(* Logix 5000 project; controller FV vendor 1 type 14 code 217 rev 31.11; software revision 31.00; part 60 of 63 *)
(* tags used below, declared in another part *)
   YP_B103 : INT[15];   // Original N File From SLC, No Description Available
   YP_B103_1_1_Storagebit : BOOL;
   YP_B30 : INT[37];   // Original N File From SLC, No Description Available
   YP_B31 : INT[37];   // Original N File From SLC, No Description Available
   YP_B92 : INT[105];   // Original N File From SLC, No Description Available
   YP_N32 : INT[257];
   YP_N55 : INT[244];   // Original N File From SLC, No Description Available
   YP_N7 : INT[56];   // INTEGER
   YP_SYSTEM_4_BIT6_TIMEBASE : ALIAS FOR One_Second_1_scan;
(* YP_Common, continued *)

   47: [AND(YP_B92[4],YP_B92[44],YP_B92[44]) ,OR(YP_B92[4],YP_B92[24],YP_B92[64]) ,XOR(YP_B92[44],YP_B92[64],YP_B92[24]) ];
   48: [AND(YP_B92[5],YP_B92[45],YP_B92[45]) ,OR(YP_B92[5],YP_B92[25],YP_B92[65]) ,XOR(YP_B92[45],YP_B92[65],YP_B92[25]) ];
   49: [AND(YP_B92[6],YP_B92[46],YP_B92[46]) ,OR(YP_B92[6],YP_B92[26],YP_B92[66]) ,XOR(YP_B92[46],YP_B92[66],YP_B92[26]) ];
   50: [AND(YP_B92[7],YP_B92[47],YP_B92[47]) ,OR(YP_B92[7],YP_B92[27],YP_B92[67]) ,XOR(YP_B92[47],YP_B92[67],YP_B92[27]) ];
   51: [AND(YP_B92[8],YP_B92[48],YP_B92[48]) ,OR(YP_B92[8],YP_B92[28],YP_B92[68]) ,XOR(YP_B92[48],YP_B92[68],YP_B92[28]) ];
   52: [AND(YP_B92[9],YP_B92[49],YP_B92[49]) ,OR(YP_B92[9],YP_B92[29],YP_B92[69]) ,XOR(YP_B92[49],YP_B92[69],YP_B92[29]) ];
   53: [AND(YP_B92[10],YP_B92[50],YP_B92[50]) ,OR(YP_B92[10],YP_B92[30],YP_B92[70]) ,XOR(YP_B92[50],YP_B92[70],YP_B92[30]) ];
   54: [AND(YP_B92[11],YP_B92[51],YP_B92[51]) ,OR(YP_B92[11],YP_B92[31],YP_B92[71]) ,XOR(YP_B92[51],YP_B92[71],YP_B92[31]) ];
   55: [AND(YP_B92[12],YP_B92[52],YP_B92[52]) ,OR(YP_B92[12],YP_B92[32],YP_B92[72]) ,XOR(YP_B92[52],YP_B92[72],YP_B92[32]) ];
   56: [AND(YP_B92[13],YP_B92[53],YP_B92[53]) ,OR(YP_B92[13],YP_B92[33],YP_B92[73]) ,XOR(YP_B92[53],YP_B92[73],YP_B92[33]) ];
   57: [AND(YP_B92[14],YP_B92[54],YP_B92[54]) ,OR(YP_B92[14],YP_B92[34],YP_B92[74]) ,XOR(YP_B92[54],YP_B92[74],YP_B92[34]) ];
   58: [AND(YP_B92[15],YP_B92[55],YP_B92[55]) ,OR(YP_B92[15],YP_B92[35],YP_B92[75]) ,XOR(YP_B92[55],YP_B92[75],YP_B92[35]) ];
   59: [AND(YP_B92[16],YP_B92[56],YP_B92[56]) ,OR(YP_B92[16],YP_B92[36],YP_B92[76]) ,XOR(YP_B92[56],YP_B92[76],YP_B92[36]) ];
   60: [AND(YP_B92[17],YP_B92[57],YP_B92[57]) ,OR(YP_B92[17],YP_B92[37],YP_B92[77]) ,XOR(YP_B92[57],YP_B92[77],YP_B92[37]) ];
   61: [AND(YP_B92[18],YP_B92[58],YP_B92[58]) ,OR(YP_B92[18],YP_B92[38],YP_B92[78]) ,XOR(YP_B92[58],YP_B92[78],YP_B92[38]) ];
   62: [AND(YP_B92[19],YP_B92[59],YP_B92[59]) ,OR(YP_B92[19],YP_B92[39],YP_B92[79]) ,XOR(YP_B92[59],YP_B92[79],YP_B92[39]) ];
   63: [XIC(YP_B30[31].4) ,XIC(YP_B103[1].2) ]OSR(YP_B103[1].1,YP_B103_1_1_Storagebit)XIC(YP_B103_1_1_Storagebit)OTE(YP_B103[1].0);
   64: XIC(YP_B103[1].2)OTU(YP_B103[1].2);
   65: XIC(YP_B103[1].0)[OR(YP_B92[20],YP_B92[40],YP_B92[40]) ,AND(YP_B92[0],YP_B92[20],YP_B92[20]) ];
   66: XIC(YP_B103[1].0)[OR(YP_B92[21],YP_B92[41],YP_B92[41]) ,AND(YP_B92[1],YP_B92[21],YP_B92[21]) ];
   67: XIC(YP_B103[1].0)[OR(YP_B92[22],YP_B92[42],YP_B92[42]) ,AND(YP_B92[2],YP_B92[22],YP_B92[22]) ];
   68: XIC(YP_B103[1].0)[OR(YP_B92[23],YP_B92[43],YP_B92[43]) ,AND(YP_B92[3],YP_B92[23],YP_B92[23]) ];
   69: XIC(YP_B103[1].0)[OR(YP_B92[24],YP_B92[44],YP_B92[44]) ,AND(YP_B92[4],YP_B92[24],YP_B92[24]) ];
   70: XIC(YP_B103[1].0)[OR(YP_B92[25],YP_B92[45],YP_B92[45]) ,AND(YP_B92[5],YP_B92[25],YP_B92[25]) ];
   71: XIC(YP_B103[1].0)[OR(YP_B92[26],YP_B92[46],YP_B92[46]) ,AND(YP_B92[6],YP_B92[26],YP_B92[26]) ];
   72: XIC(YP_B103[1].0)[OR(YP_B92[27],YP_B92[47],YP_B92[47]) ,AND(YP_B92[7],YP_B92[27],YP_B92[27]) ];
   73: XIC(YP_B103[1].0)[OR(YP_B92[28],YP_B92[48],YP_B92[48]) ,AND(YP_B92[8],YP_B92[28],YP_B92[28]) ];
   74: XIC(YP_B103[1].0)[OR(YP_B92[29],YP_B92[49],YP_B92[49]) ,AND(YP_B92[9],YP_B92[29],YP_B92[29]) ];
   75: XIC(YP_B103[1].0)[OR(YP_B92[30],YP_B92[50],YP_B92[50]) ,AND(YP_B92[10],YP_B92[30],YP_B92[30]) ];
   76: XIC(YP_B103[1].0)[OR(YP_B92[31],YP_B92[51],YP_B92[51]) ,AND(YP_B92[11],YP_B92[31],YP_B92[31]) ];
   77: XIC(YP_B103[1].0)[OR(YP_B92[32],YP_B92[52],YP_B92[52]) ,AND(YP_B92[12],YP_B92[32],YP_B92[32]) ];
   78: XIC(YP_B103[1].0)[OR(YP_B92[33],YP_B92[53],YP_B92[53]) ,AND(YP_B92[13],YP_B92[33],YP_B92[33]) ];
   79: XIC(YP_B103[1].0)[OR(YP_B92[34],YP_B92[54],YP_B92[54]) ,AND(YP_B92[14],YP_B92[34],YP_B92[34]) ];
   80: XIC(YP_B103[1].0)[OR(YP_B92[35],YP_B92[55],YP_B92[55]) ,AND(YP_B92[15],YP_B92[35],YP_B92[35]) ];
   81: XIC(YP_B103[1].0)[OR(YP_B92[36],YP_B92[56],YP_B92[56]) ,AND(YP_B92[16],YP_B92[36],YP_B92[36]) ];
   82: XIC(YP_B103[1].0)[OR(YP_B92[37],YP_B92[57],YP_B92[57]) ,AND(YP_B92[17],YP_B92[37],YP_B92[37]) ];
   83: XIC(YP_B103[1].0)[OR(YP_B92[38],YP_B92[58],YP_B92[58]) ,AND(YP_B92[18],YP_B92[38],YP_B92[38]) ];
   84: XIC(YP_B103[1].0)[OR(YP_B92[39],YP_B92[59],YP_B92[59]) ,AND(YP_B92[19],YP_B92[39],YP_B92[39]) ];
   85: XIC(YP_B103[1].0)MOV(0,YP_N7[38]);
   86: XIC(YP_SYSTEM_4_BIT6_TIMEBASE)MOV(YP_B92[60],YP_B92[80]);
   87: XIO(YP_SYSTEM_4_BIT6_TIMEBASE)MOV(YP_B92[40],YP_B92[80]);
   88: XIC(YP_SYSTEM_4_BIT6_TIMEBASE)MOV(YP_B92[61],YP_B92[81]);
   89: XIO(YP_SYSTEM_4_BIT6_TIMEBASE)MOV(YP_B92[41],YP_B92[81]);
   90: XIC(YP_SYSTEM_4_BIT6_TIMEBASE)MOV(YP_B92[62],YP_B92[82]);
   91: XIO(YP_SYSTEM_4_BIT6_TIMEBASE)MOV(YP_B92[42],YP_B92[82]);
   92: XIC(YP_SYSTEM_4_BIT6_TIMEBASE)MOV(YP_B92[63],YP_B92[83]);
   93: XIO(YP_SYSTEM_4_BIT6_TIMEBASE)MOV(YP_B92[43],YP_B92[83]);
   94: XIC(YP_SYSTEM_4_BIT6_TIMEBASE)MOV(YP_B92[64],YP_B92[84]);
   95: XIO(YP_SYSTEM_4_BIT6_TIMEBASE)MOV(YP_B92[44],YP_B92[84]);
   96: XIC(YP_SYSTEM_4_BIT6_TIMEBASE)MOV(YP_B92[65],YP_B92[85]);
   97: XIO(YP_SYSTEM_4_BIT6_TIMEBASE)MOV(YP_B92[45],YP_B92[85]);
   98: XIC(YP_SYSTEM_4_BIT6_TIMEBASE)MOV(YP_B92[66],YP_B92[86]);
   99: XIO(YP_SYSTEM_4_BIT6_TIMEBASE)MOV(YP_B92[46],YP_B92[86]);
   100: XIC(YP_SYSTEM_4_BIT6_TIMEBASE)MOV(YP_B92[67],YP_B92[87]);
   101: XIO(YP_SYSTEM_4_BIT6_TIMEBASE)MOV(YP_B92[47],YP_B92[87]);
   102: XIC(YP_SYSTEM_4_BIT6_TIMEBASE)MOV(YP_B92[68],YP_B92[88]);
   103: XIO(YP_SYSTEM_4_BIT6_TIMEBASE)MOV(YP_B92[48],YP_B92[88]);
   104: XIC(YP_SYSTEM_4_BIT6_TIMEBASE)MOV(YP_B92[69],YP_B92[89]);
   105: XIO(YP_SYSTEM_4_BIT6_TIMEBASE)MOV(YP_B92[49],YP_B92[89]);
   106: XIC(YP_SYSTEM_4_BIT6_TIMEBASE)MOV(YP_B92[70],YP_B92[90]);
   107: XIO(YP_SYSTEM_4_BIT6_TIMEBASE)MOV(YP_B92[50],YP_B92[90]);
   108: XIC(YP_SYSTEM_4_BIT6_TIMEBASE)MOV(YP_B92[71],YP_B92[91]);
   109: XIO(YP_SYSTEM_4_BIT6_TIMEBASE)MOV(YP_B92[51],YP_B92[91]);
   110: XIC(YP_SYSTEM_4_BIT6_TIMEBASE)MOV(YP_B92[72],YP_B92[92]);
   111: XIO(YP_SYSTEM_4_BIT6_TIMEBASE)MOV(YP_B92[52],YP_B92[92]);
   112: XIC(YP_SYSTEM_4_BIT6_TIMEBASE)MOV(YP_B92[73],YP_B92[93]);
   113: XIO(YP_SYSTEM_4_BIT6_TIMEBASE)MOV(YP_B92[53],YP_B92[93]);
   114: XIC(YP_SYSTEM_4_BIT6_TIMEBASE)MOV(YP_B92[74],YP_B92[94]);
   115: XIO(YP_SYSTEM_4_BIT6_TIMEBASE)MOV(YP_B92[54],YP_B92[94]);
   116: XIC(YP_SYSTEM_4_BIT6_TIMEBASE)MOV(YP_B92[75],YP_B92[95]);
   117: XIO(YP_SYSTEM_4_BIT6_TIMEBASE)MOV(YP_B92[55],YP_B92[95]);
   118: XIC(YP_SYSTEM_4_BIT6_TIMEBASE)MOV(YP_B92[76],YP_B92[96]);
   119: XIO(YP_SYSTEM_4_BIT6_TIMEBASE)MOV(YP_B92[56],YP_B92[96]);
   120: XIC(YP_SYSTEM_4_BIT6_TIMEBASE)MOV(YP_B92[77],YP_B92[97]);
   121: XIO(YP_SYSTEM_4_BIT6_TIMEBASE)MOV(YP_B92[57],YP_B92[97]);
   122: XIC(YP_SYSTEM_4_BIT6_TIMEBASE)MOV(YP_B92[78],YP_B92[98]);
   123: XIO(YP_SYSTEM_4_BIT6_TIMEBASE)MOV(YP_B92[58],YP_B92[98]);
   124: XIC(YP_SYSTEM_4_BIT6_TIMEBASE)MOV(YP_B92[79],YP_B92[99]);
   125: XIO(YP_SYSTEM_4_BIT6_TIMEBASE)MOV(YP_B92[59],YP_B92[99]);
   126: [NEQ(YP_B92[20],0) ,NEQ(YP_B92[21],0) ,NEQ(YP_B92[22],0) ,NEQ(YP_B92[23],0) ,NEQ(YP_B92[24],0) ,NEQ(YP_B92[25],0) ,NEQ(YP_B92[26],0) ,NEQ(YP_B92[27],0) ,NEQ(YP_B92[28],0) ,NEQ(YP_B92[29],0) ,NEQ(YP_B92[30],0) ,NEQ(YP_B92[31],0) ,NEQ(YP_B92[32],0) ,NEQ(YP_B92[33],0) ,NEQ(YP_B92[34],0) ,NEQ(YP_B92[35],0) ,NEQ(YP_B92[36],0) ,NEQ(YP_B92[37],0) ,NEQ(YP_B92[38],0) ,NEQ(YP_B92[39],0) ]OTE(YP_B31[31].4);
   127: MOV(YP_B92[0],YP_N55[219])MOV(YP_B92[1],YP_N55[220]);
   128: MOV(YP_B92[0],YP_N32[219])MOV(YP_B92[1],YP_N32[220]);
END_ROUTINE
